// Mitsubishi GX Works2 project: 20国轩1次注液出11.16和条码枪通信   PLC: Q06UDEH (continued)
	
	(*U1任务处理 *)
	m_TPU1TaskComplete(IN:=ConveyorIO20110.xEmpty ,PT:=t#200ms,Q:= m_xU1TaskComplete,ET:= m_tU1TaskComplete );
	(*这里东西运走之后延时200ms再完成任务，这个时间是防止扫描周期的影响，让U型块先复位，再完成任务*)
Task20301(	xCondition:=TaskCondition20301,
 xTaskComplete:=LDF(TRUE,m_xU1TaskComplete),
 xReset:=g_xResetSingle AND g_diDeviceIDSelect=20110,
 iPriority:=UConveyorIO20301.iTask);
	TaskCondition20301[1]:=NOT ConveyorIO20101.xEmpty  AND LifterIO20201.iCurrentPos=2  AND X2F AND m_i20101Task>0;
	TaskCondition20301[2]:=(NOT ConveyorIO201021.xEmpty AND ConveyorIO201021.diDesConveyor=20115) 
												OR(NOT  ConveyorIO20110.xEmpty AND (ConveyorIO20110.diDesConveyor<>20102 OR ConveyorIO20110.diDesConveyor<>20103)) ;
	TaskCondition20301[3]:=(NOT ConveyorIO201031.xEmpty AND ConveyorIO201031.diDesConveyor=20115)
												OR (NOT  ConveyorIO20110.xEmpty AND(ConveyorIO20110.diDesConveyor<>20102 OR ConveyorIO20110.diDesConveyor<>20103));
	(*U2Task	*)
	m_TPU2TaskComplete(IN:=ConveyorIO20111.xEmpty ,PT:=t#200ms,Q:= m_xU2TaskComplete,ET:= m_tU2TaskComplete );
	Task20303(	xCondition:=TaskCondition20303,
 	xTaskComplete:=LDf(TRUE, m_xU2TaskComplete),
 	xReset:=g_xResetSingle AND g_diDeviceIDSelect=20111,
 	iPriority:=UConveyorIO20303.iTask);
		TaskCondition20303[1]:=NOT ConveyorIO20110.xEmpty AND NOT  (ConveyorIO20110.diDesConveyor=20103 
																OR ConveyorIO20110.diDesConveyor=20102
																OR ConveyorIO20110.diDesConveyor=0)(*不去左，不去右，也不是0，就认为可以接料*);
		TaskCondition20303[2]:=(NOT ConveyorIO201041.xEmpty  AND ConveyorIO201041.diDesConveyor=20115) 
													OR (NOT ConveyorIO20111.xEmpty AND (ConveyorIO20111.diDesConveyor<>20103 OR ConveyorIO20111.diDesConveyor<>20102) );
		TaskCondition20303[3]:=(NOT ConveyorIO201051.xEmpty  AND ConveyorIO201051.diDesConveyor=20115) 
													OR (NOT ConveyorIO20111.xEmpty AND (ConveyorIO20111.diDesConveyor<>20103 OR ConveyorIO20111.diDesConveyor<>20102));
	(*//U3Task*)
	m_TPU3TaskComplete(IN:=ConveyorIO20113.xEmpty ,PT:=t#200ms,Q:= m_xU3TaskComplete,ET:= m_tU3TaskComplete );
	Task20305(	xCondition:=TaskCondition20305,
 	xTaskComplete:=LDF(TRUE,m_xU3TaskComplete),
 	xReset:=g_xResetSingle AND g_diDeviceIDSelect=20113,
 	iPriority:=UConveyorIO20305.iTask);
		TaskCondition20305[1]:=NOT ConveyorIO20112.xEmpty(* AND  (ConveyorIO20112.diDesConveyor=20104 
																OR ConveyorIO20112.diDesConveyor=20105
																OR ConveyorIO20112.diDesConveyor=0);(*不去左，不去右，也不是0，就认为可以接料*) ;
		TaskCondition20305[2]:=(NOT ConveyorIO201061.xEmpty AND ConveyorIO201061.diDesConveyor=20115) 
													OR (NOT ConveyorIO20113.xEmpty AND (ConveyorIO20113.diDesConveyor<>20104 OR ConveyorIO20113.diDesConveyor<>20105));
		TaskCondition20305[3]:=(NOT ConveyorIO201071.xEmpty AND ConveyorIO201071.diDesConveyor=20115)
													OR (NOT ConveyorIO20113.xEmpty AND  (ConveyorIO20113.diDesConveyor<>20104 OR ConveyorIO20113.diDesConveyor<>20105));
	(*//U4Task*)
	m_TPU4TaskComplete(IN:=ConveyorIO20114.xEmpty ,PT:=t#200ms,Q:= m_xU4TaskComplete,ET:= m_tU4TaskComplete );
	Task20307(	xCondition:=TaskCondition20307,
 	xTaskComplete:=LDF(TRUE, m_xU4TaskComplete),
 	xReset:=g_xResetSingle AND g_diDeviceIDSelect=20114,
 	iPriority:=UConveyorIO20307.iTask);
		TaskCondition20307[1]:=NOT ConveyorIO20113.xEmpty  AND NOT (ConveyorIO20113.diDesConveyor=20106
																OR ConveyorIO20113.diDesConveyor=20107
																OR ConveyorIO20113.diDesConveyor=0)
(*																AND ConveyorIo20115.xEmpty*);		
		TaskCondition20307[3]:=((NOT ConveyorIO201091.xEmpty AND ConveyorIO201091.diDesConveyor=20115)
													OR (NOT ConveyorIO20114.xEmpty AND (ConveyorIO20114.diDesConveyor<>20109 OR ConveyorIO20114.diDesConveyor<>20108) ))
(*													AND ConveyorIo20115.xEmpty*);
		TaskCondition20307[2]:=((NOT ConveyorIO201081.xEmpty AND ConveyorIO201081.diDesConveyor=20115)
													OR (NOT ConveyorIO20114.xEmpty AND (ConveyorIO20114.diDesConveyor<>20109 OR ConveyorIO20114.diDesConveyor<>20108) ))
(*													AND ConveyorIo20115.xEmpty*);
(*目标地址的传递，横纵分开传递*)
	ConveyorIO20110.diDesConveyorIn:=	ConveyorIO20101.diDesConveyorOut;
	ConveyorIO20111.diDesConveyorIn:=	ConveyorIO20110.diDesConveyorOut;
	ConveyorIO20112.diDesConveyorIn:=	ConveyorIO20111.diDesConveyorOut;
	ConveyorIO20113.diDesConveyorIn:=	ConveyorIO20112.diDesConveyorOut;
	ConveyorIO20114.diDesConveyorIn:=	ConveyorIO20113.diDesConveyorOut;		
(*纵向传递*)
	ConveyorIO20102.diDesConveyorIn:=	ConveyorIO201021.diDesConveyorOut;
	ConveyorIO20103.diDesConveyorIn:=	ConveyorIO201031.diDesConveyorOut;
	ConveyorIO20104.diDesConveyorIn:=	ConveyorIO201041.diDesConveyorOut;
	ConveyorIO20105.diDesConveyorIn:=	ConveyorIO201051.diDesConveyorOut;
	ConveyorIO20106.diDesConveyorIn:=	ConveyorIO201061.diDesConveyorOut;
	ConveyorIO20107.diDesConveyorIn:=	ConveyorIO201071.diDesConveyorOut;
	ConveyorIO20108.diDesConveyorIn:=	ConveyorIO201081.diDesConveyorOut;
	ConveyorIO20109.diDesConveyorIn:=	ConveyorIO201091.diDesConveyorOut;	
	

IF g_xAuto THEN
	D201.0:=ConveyorIO201221.xEmpty;
	Switchio20311.xEntryEnable:=
	D401.0;(*两个PLC通信，以太网方式*)
	Switchio20311.xSwithEnable:=1;
	Switchio20311.xExitEnable:=ConveyorIO201231.xEmpty;
	ConveyorIO201231.xLoad:=ConveyorIO20122.xNextRun;
	ConveyorIO201231.xUnload:=ConveyorIO20123.xEmpty;
	ConveyorIO20123.xLoad:=	ConveyorIO201231.xNextRun;;	
	ConveyorIO20123.xUnload:=	ConveyorIO20124.xEmpty;
	ConveyorIO20124.xLoad:=	ConveyorIO20123.xNextRun;	
	ConveyorIO20124.xUnload:=	ConveyorIO20125.xEmpty;
	SwitchIO20312.xEntryEnable:=ConveyorIO20124.xNextRun;
	SwitchIO20312.xSwithEnable:=1;
	SwitchIO20312.xLiftCylinderExtendInit:=1;
	SwitchIO20312.xExitEnable:=ConveyorIO201261.xEmpty;     
	ConveyorIO201261.xLoad:=ConveyorIO20126.xNextRun;
	ConveyorIO201261.xUnload:=ConveyorIO20127.xEmpty;
	ConveyorIO20127.xLoad:=	ConveyorIO201261.xNextRun;	
	ConveyorIO20127.xUnload:=	ConveyorIO20128.xEmpty;
	ConveyorIO20128.xLoad:=	ConveyorIO20127.xNextRun;	
	ConveyorIO20128.xUnload:=	ConveyorIO20129.xEmpty;
	ConveyorIO20129.xLoad:=	ConveyorIO20128.xNextRun;	
	ConveyorIO20129.xUnload:=	ConveyorIO20130.xEmpty AND NOT ConveyorIO20130.xError;
	ConveyorIO20130.xLoad:=	ConveyorIO20129.xNextRun;	
	ConveyorIO20130.xUnload:=ConveyorIO20101.xEmpty AND LifterIO20201.iCurrentPos=1 AND X2E AND NOT ConveyorIO20101.xError;
	ConveyorIO20101.xLoad:=ConveyorIO20130.xNextRun AND LifterIO20201.iCurrentPos=1 AND X2E;(*运到升降机上了*)
	LifterIO20201.xMDIExe:=NOT 	ConveyorIO20101.xError
													AND NOT ConveyorIO20130.xError
													AND NOT ConveyorIO20110.xError;
	IF ConveyorIO20101.xEmpty THEN
		LifterIO20201.iDestinationPos:=1;
	ELSE
		LifterIO20201.iDestinationPos:=2;
	END_IF;
	m_TonU1TaskStart(IN:=ConveyorIO20110.xEmpty AND UConveyorIO20301.iTask=1  ,PT:= t#1s ,Q:=m_xU1TaskStart,ET:= m_tU1TaskStart );
	ConveyorIO20101.xUnload:=m_xU1TaskStart  AND 
   															LifterIO20201.iCurrentPos=2 AND X2F
 															 (*AND UConveyorIO20301.iTask=1       这个信号会波动
 															 AND ConveyorIO20110.xEmpty*);
 	ConveyorIO20101.xUnloadCCW:=1;
   
	(*//U1*)	
	UConveyorIO20301.xEntryEnable1:= ConveyorIO20101.xNextRun;
	UConveyorIO20301.xEntryEnable2:=ConveyorIO201021.xNextRun;
	UConveyorIO20301.xEntryEnable3:=ConveyorIO201031.xNextRun;
	
	m_TonU2TaskStart(IN:=ConveyorIO20111.xEmpty  ,PT:= t#300ms ,Q:=m_xU2TaskStart,ET:= m_tU2TaskStart );
	UConveyorIO20301.xExitEnable1:= m_xU2TaskStart AND UConveyorIO20303.iTask=1;
	UConveyorIO20301.xExitEnable2:=ConveyorIO201021.xEmpty;
	UConveyorIO20301.xExitEnable3:=ConveyorIO201031.xEmpty;
	(*//U1接料*)
	ConveyorIO201021.xload:=	ConveyorIO20102.xNextRun;
	ConveyorIO201031.xload:=	ConveyorIO20103.xNextRun;
	(*单电控夹紧气缸动作控制*)
	m_xCatchCylinder[2]:=NOT ConveyorIO201021.xEmpty AND ConveyorIO201021.diDesConveyor=0;
	m_xCatchCylinder[3]:=NOT ConveyorIO201031.xEmpty AND ConveyorIO201031.diDesConveyor=0;
	(*//U1出料Unload	*)
		ConveyorIO201021.xUnload:=ConveyorIO20102.xEmpty AND UConveyorIO20301.iTask=2;
		ConveyorIO201031.xUnload:=ConveyorIO20103.xEmpty AND UConveyorIO20301.iTask=3;

	(**//U2*)
	UConveyorIO20303.xEntryEnable1:= ConveyorIO20110.xNextRun ;
	UConveyorIO20303.xEntryEnable2:=ConveyorIO201041.xNextRun;
	UConveyorIO20303.xEntryEnable3:=ConveyorIO201051.xNextRun;
	UConveyorIO20303.xExitEnable1:= ConveyorIO20112.xEmpty;
	UConveyorIO20303.xExitEnable2:=ConveyorIO201041.xEmpty;
	UConveyorIO20303.xExitEnable3:=ConveyorIO201051.xEmpty;
	(*//U2接料	*)
	ConveyorIO201041.xload:=	ConveyorIO20104.xNextRun;
	ConveyorIO201051.xload:=	ConveyorIO20105.xNextRun;
		(*单电控夹紧气缸动作控制*)
	m_xCatchCylinder[4]:=NOT ConveyorIO201041.xEmpty AND ConveyorIO201041.diDesConveyor=0;
	m_xCatchCylinder[5]:=NOT ConveyorIO201051.xEmpty AND ConveyorIO201051.diDesConveyor=0;
	(*//U2出料Unload	*)
		ConveyorIO201041.xUnload:=ConveyorIO20104.xEmpty AND UConveyorIO20303.iTask=2;
		ConveyorIO201051.xUnload:=ConveyorIO20105.xEmpty AND UConveyorIO20303.iTask=3;
	(*//中间传输*)
	ConveyorIO20112.xLoad:=ConveyorIO20111.xNextRun;
	m_TonU3TaskStart(IN:=ConveyorIO20113.xEmpty  ,PT:= t#300ms ,Q:=m_xU3TaskStart,ET:= m_tU3TaskStart );
	ConveyorIO20112.xUnload:=m_xU3TaskStart AND UConveyorIO20305.iTask=1;
	
	(*//U3	*)
	UConveyorIO20305.xEntryEnable1:= ConveyorIO20112.xNextRun;
	UConveyorIO20305.xEntryEnable2:=ConveyorIO201061.xNextRun;
	UConveyorIO20305.xEntryEnable3:=ConveyorIO201071.xNextRun;
	
	m_TonU4TaskStart(IN:=ConveyorIO20114.xEmpty  ,PT:= t#300ms ,Q:=m_xU4TaskStart,ET:= m_tU4TaskStart );
	UConveyorIO20305.xExitEnable1:= m_xU4TaskStart AND UConveyorIO20307.iTask=1 ;
	UConveyorIO20305.xExitEnable2:=ConveyorIO201061.xEmpty;
	UConveyorIO20305.xExitEnable3:=ConveyorIO201071.xEmpty;
	(*	//U3接料*)
	ConveyorIO201061.xload:=	ConveyorIO20106.xNextRun;
	ConveyorIO201071.xload:=	ConveyorIO20107.xNextRun;
		(*单电控夹紧气缸动作控制*)
	m_xCatchCylinder[6]:=NOT ConveyorIO201061.xEmpty AND ConveyorIO201061.diDesConveyor=0;
	m_xCatchCylinder[7]:=NOT ConveyorIO201071.xEmpty AND ConveyorIO201071.diDesConveyor=0;
	(*//U3出料Unload	*)
		ConveyorIO201061.xUnload:=ConveyorIO20106.xEmpty AND  UConveyorIO20305.iTask=2;
		ConveyorIO201071.xUnload:=ConveyorIO20107.xEmpty AND UConveyorIO20305.iTask=3;
	
	(*//U4	*)
	UConveyorIO20307.xEntryEnable1:= ConveyorIO20113.xNextRun ;
	UConveyorIO20307.xEntryEnable2:=ConveyorIO201081.xNextRun;
	UConveyorIO20307.xEntryEnable3:=ConveyorIO201091.xNextRun;
	UConveyorIO20307.xExitEnable1:= ConveyorIO20115.xEmpty ;
	UConveyorIO20307.xExitEnable2:=ConveyorIO201081.xEmpty;
	UConveyorIO20307.xExitEnable3:=ConveyorIO201091.xEmpty;
	(*	//U4接料*)
	ConveyorIO201081.xload:=	ConveyorIO20108.xNextRun;
	ConveyorIO201091.xload:=	ConveyorIO20109.xNextRun;
		(*单电控夹紧气缸动作控制*)
	m_xCatchCylinder[8]:=NOT ConveyorIO201081.xEmpty AND ConveyorIO201081.diDesConveyor=0;
	m_xCatchCylinder[9]:=NOT ConveyorIO201091.xEmpty AND ConveyorIO201091.diDesConveyor=0;
	(*//U4出料Unload	*)
	ConveyorIO201081.xUnload:=ConveyorIO20108.xEmpty AND UConveyorIO20307.iTask=2;
	ConveyorIO201091.xUnload:=ConveyorIO20109.xEmpty AND UConveyorIO20307.iTask=3;
	SwitchIO20309.xEntryEnable:=	ConveyorIO20114.xNextRun;
	SwitchIO20309.xSwithEnable:=1;
	SwitchIO20309.xExitEnable:=ConveyorIO201161.xEmpty;
	ConveyorIO201161.xLoad:=ConveyorIO20116.xNextRun;
	ConveyorIO201161.xUnload:=ConveyorIO20117.xEmpty;
	ConveyorIO20117.xLoad:=ConveyorIO201161.xNextRun;
	ConveyorIO20117.xUnload:=ConveyorIO20118.xEmpty;
	ConveyorIO20118.xLoad:=ConveyorIO20117.xNextRun;
	ConveyorIO20118.xUnload:=ConveyorIO20119.xEmpty AND (g_xScanDone OR SM400);
	Y252:=NOT ConveyorIO20118.xNextRun;
	ConveyorIo20119.tLoadDelay:=T#6s;	
	SwitchIO20310.xEntryEnable:=ConveyorIO20118.xNextRun;
	SwitchIO20310.xLiftCylinderExtendInit:=1;
	SwitchIO20310.xSwithEnable:=1;
	SwitchIO20310.xExitEnable:=D401.2;
	D201.2:=ConveyorIO201191.xNextRun;
(*	ConveyorIO20119.xPutInto:=NOT ConveyorIO20119.xCWPresent AND SM412;
	ConveyorIO201191.xPutInto:=NOT ConveyorIO201191.xCWPresent AND SM412;*)
	(*至此，托盘循环完成*)
	
END_IF;(*g_xAuto那个IF**)	
	(*******************************以下部分为机械手控制*********************************************)
		(*1号机器人*)
		(*位置1*)
		(*发送给机器人的可以放料信号*)
	g_xRobot1Pos1Ready:=NOT ConveyorIO201021.xEmpty   (*线体不为空*)
												AND ConveyorIO201021.diDesConveyor=0(*无目标线体位置*)
												AND NOT g_xRobot1Pos2Ready(*与位置2的信号互锁，同时只有一个ready信号*)
												AND g_xAuto;
		(*接收机器人的完成信号*)
	DMOV(g_xRobot1Pos1Done,20115,ConveyorIO201021.diDesConveyor);(*将目标位置设置成出料线体*)
		(*位置2*)
		(*发送给机器人的可以放料信号*)
	g_xRobot1Pos2Ready:=NOT ConveyorIO201031.xEmpty  (*线体不为空*)
												AND ConveyorIO201031.diDesConveyor=0(*无目标线体位置*)
												AND NOT g_xRobot1Pos1Ready(*与位置1的信号互锁，同时只有一个ready信号*)
												AND g_xAuto;
			(*接收机器人的完成信号*)
	DMOV(g_xRobot1Pos2Done,20115,ConveyorIO201031.diDesConveyor);
	(*2号机器人*)
	g_xRobot2Pos1Ready:=NOT ConveyorIO201041.xEmpty 
												AND ConveyorIO201041.diDesConveyor=0
												AND NOT g_xRobot2Pos2Ready
												AND g_xAuto;
	DMOV(g_xRobot2Pos1Done,20115,ConveyorIO201041.diDesConveyor);
	g_xRobot2Pos2Ready:=NOT ConveyorIO201051.xEmpty 
												AND ConveyorIO201051.diDesConveyor=0
												AND NOT g_xRobot2Pos1Ready 
												AND g_xAuto;
	DMOV(g_xRobot2Pos2Done,20115,ConveyorIO201051.diDesConveyor);
			(*3号机器人*)
		(*位置1*)
		(*发送给机器人的可以放料信号*)
	g_xRobot3Pos1Ready:=NOT ConveyorIO201061.xEmpty   (*线体不为空*)
												AND ConveyorIO201061.diDesConveyor=0(*无目标线体位置*)
												AND NOT g_xRobot3Pos2Ready(*与位置2的信号互锁，同时只有一个ready信号*)
												AND g_xAuto;
		(*接收机器人的完成信号*)
	DMOV(g_xRobot3Pos1Done,20115,ConveyorIO201061.diDesConveyor);(*将目标位置设置成出料线体*)
		(*位置2*)
		(*发送给机器人的可以放料信号*)
	g_xRobot3Pos2Ready:=NOT ConveyorIO201071.xEmpty  (*线体不为空*)
												AND ConveyorIO201071.diDesConveyor=0(*无目标线体位置*)
												AND NOT g_xRobot3Pos1Ready(*与位置1的信号互锁，同时只有一个ready信号*) 
												AND g_xAuto;
			(*接收机器人的完成信号*)
	DMOV(g_xRobot3Pos2Done,20115,ConveyorIO201071.diDesConveyor);
			(*4号机器人*)
		(*位置1*)
		(*发送给机器人的可以放料信号*)
	g_xRobot4Pos1Ready:=NOT ConveyorIO201081.xEmpty   (*线体不为空*)
												AND ConveyorIO201081.diDesConveyor=0(*无目标线体位置*)
												AND NOT g_xRobot4Pos2Ready(*与位置2的信号互锁，同时只有一个ready信号*) 
												AND g_xAuto;
		(*接收机器人的完成信号*)
	DMOV(g_xRobot4Pos1Done,20115,ConveyorIO201081.diDesConveyor);(*将目标位置设置成出料线体*)
		(*位置4*)
		(*发送给机器人的可以放料信号*)
	g_xRobot4Pos2Ready:=NOT ConveyorIO201091.xEmpty  (*线体不为空*)
												AND ConveyorIO201091.diDesConveyor=0(*无目标线体位置*)
												AND NOT g_xRobot4Pos1Ready(*与位置1的信号互锁，同时只有一个ready信号*) 
												AND g_xAuto;
			(*接收机器人的完成信号*)
	DMOV(g_xRobot4Pos2Done,20115,ConveyorIO201091.diDesConveyor);
		
	(*******************************以上部分为机械手控制*********************************************)
	
IF NOT g_xAuto THEN
	D201.0:=0;
	D201.2:=0;
	ConveyorIO201021.diDesConveyor:=0;
	ConveyorIO201031.diDesConveyor:=0;	
	ConveyorIO201041.diDesConveyor:=0;
	ConveyorIO201051.diDesConveyor:=0;
	ConveyorIO201061.diDesConveyor:=0;
	ConveyorIO201071.diDesConveyor:=0;	
	ConveyorIO201081.diDesConveyor:=0;
	ConveyorIO201091.diDesConveyor:=0;	
	g_xRobot1Pos1Ready:=0;
	g_xRobot1Pos2Ready:=0;
	g_xRobot2Pos1Ready:=0;
	g_xRobot2Pos2Ready:=0;
	g_xRobot3Pos1Ready:=0;
	g_xRobot3Pos2Ready:=0;
	g_xRobot4Pos1Ready:=0;
	g_xRobot4Pos2Ready:=0;
	
END_IF;
(*//统计计数*)

ADD_E(LDP(TRUE,NOT ConveyorIO201021.xEmpty)AND UConveyorIO20301.iTask=1,	D10,	1,	D10 );
ADD_E(LDP(TRUE,NOT ConveyorIO201031.xEmpty)AND UConveyorIO20301.iTask=1,	D12,	1,	D12 );
ADD_E(LDP(TRUE,NOT ConveyorIO201041.xEmpty)AND UConveyorIO20303.iTask=1,	D14,	1,	D14 );
ADD_E(LDP(TRUE,NOT ConveyorIO201051.xEmpty)AND UConveyorIO20303.iTask=1,	D16,	1,	D16 );
ADD_E(LDP(TRUE,NOT ConveyorIO201061.xEmpty)AND UConveyorIO20305.iTask=1,	D18,	1,	D18 );
ADD_E(LDP(TRUE,NOT ConveyorIO201071.xEmpty)AND UConveyorIO20305.iTask=1,	D20,	1,	D20 );
ADD_E(LDP(TRUE,NOT ConveyorIO201081.xEmpty)AND UConveyorIO20307.iTask=1,	D22,	1,	D22 );
ADD_E(LDP(TRUE,NOT ConveyorIO201091.xEmpty)AND UConveyorIO20307.iTask=1,	D24,	1,	D24 );
(*//统计数据清零,这些M都是在触摸屏上的数据清零按钮*)
DMOV(	M62,	0,	D10);
DMOV(	M63,	0,	D12 );
DMOV(	M64,	0,	D14 );
DMOV(	M65,	0,	D16 );
DMOV(	M66,	0,	D18 );
DMOV(	M67,	0,	D20 );
DMOV(	M68,	0,	D22 );
DMOV(	M69,	0,	D24 );
(*临时加一些送出按钮，方便操作*)
DMOVP( M42 ,10115 , ConveyorIO201021.diDesConveyor );
DMOVP( M43 ,10115 , ConveyorIO201031.diDesConveyor );
DMOVP( M44 ,10115 , ConveyorIO201041.diDesConveyor );
DMOVP( M45 ,10115 , ConveyorIO201051.diDesConveyor );
DMOVP( M46 ,10115 , ConveyorIO201061.diDesConveyor );
DMOVP( M47 ,10115 , ConveyorIO201071.diDesConveyor );
DMOVP( M48 ,10115 , ConveyorIO201081.diDesConveyor );
DMOVP( M49 ,10115 , ConveyorIO201091.diDesConveyor );

(*报警*)
g_xAlarm:=NOT g_xEStop;
END_PROGRAM

FUNCTION_BLOCK PreemptivePriority
VAR_INPUT
  xCondition : ARRAY [1..13] OF BOOL;  (* 条件1 *)
  xTaskComplete : BOOL;  (* 任务完成 *)
  xReset : BOOL;  (* 复位 *)
END_VAR
VAR
  xOccupy : BOOL;  (* 占用 *)
END_VAR
VAR_OUTPUT
  iPriority : INT;  (* 输出任务号 *)
END_VAR
VAR
  m_tonConditionDelay : TON;
  m_xConditionDelay : BOOL;
  m_tConditionCurrentTime : TIME;
  m_iLastTask : INT;  (* 上次执行的任务 *)
  m_tpLastTaskPulse1 : TP;
  m_tpLastTaskPulse2 : TP;
  m_tpLastTaskPulse3 : TP;
  m_tpLastTaskPulse4 : TP;
  m_tpLastTaskPulse5 : TP;
  m_xLastTaskPulse : ARRAY [1..13] OF BOOL;
  m_tLastTaskPulse : ARRAY [1..13] OF TIME := [13(T#0s)];
  m_tpLastTaskPulse6 : TON;
  ii : INT;
END_VAR
VAR CONSTANT
  CONDITION_QUANTITY : INT := 9;
END_VAR
VAR
  m_tpLastTaskPulse7 : TON;
  m_tpLastTaskPulse8 : TON;
  m_tpLastTaskPulse9 : TON;
  m_tpLastTaskPulse10 : TON;
  m_tpLastTaskPulse11 : TON;
  m_tpLastTaskPulse12 : TON;
  m_tpLastTaskPulse13 : TON;
END_VAR
(*抢占式优先级块
现在满足13个条件的任务进行抢占式优先级排列
条件满足后延时两秒，开始执行任务，
同一任务连续执行优先级下降
需要改造成任意多个
使用于一个入口多个出口的程序，使用抢占式优先级块
*)
IF LDP(TRUE, xTaskComplete) THEN
	xOccupy:=0;
	iPriority:=0;
END_IF;
(*//任务滤波，延时两秒*)
m_tonConditionDelay(IN:=( xCondition[1]
 	OR xCondition[2]
 	OR xCondition[3]
 	OR xCondition[4]
 	OR xCondition[5]
 	OR xCondition[6]
 	OR xCondition[7]
 	OR xCondition[8]
 	OR xCondition[9]
 	OR xCondition[10]
 	OR xCondition[11]
 	OR xCondition[12]
 	OR xCondition[13]
 	)
 	AND iPriority=0,
 PT:= T#1s,
 Q:= m_xConditionDelay ,
 ET:= m_tConditionCurrentTime );		
(*//判断优先级，上个任务与本次任务相同，延时一秒执行*)
m_tpLastTaskPulse1(IN:= xCondition[1]  AND m_iLastTask=1 AND m_xConditionDelay  ,PT:= T#1s,Q:= m_xLastTaskPulse[1],ET:= m_tLastTaskPulse[1] );
m_tpLastTaskPulse2(IN:= xCondition[2]  AND m_iLastTask=2 AND m_xConditionDelay  ,PT:= T#1s,Q:= m_xLastTaskPulse[2],ET:= m_tLastTaskPulse[2] );
m_tpLastTaskPulse3(IN:= xCondition[3]  AND m_iLastTask=3 AND m_xConditionDelay  ,PT:= T#1s,Q:= m_xLastTaskPulse[3],ET:= m_tLastTaskPulse[3] );
m_tpLastTaskPulse4(IN:= xCondition[4]  AND m_iLastTask=4 AND m_xConditionDelay  ,PT:= T#1s,Q:= m_xLastTaskPulse[4],ET:= m_tLastTaskPulse[4] );
m_tpLastTaskPulse5(IN:= xCondition[5]  AND m_iLastTask=5 AND m_xConditionDelay  ,PT:= T#1s,Q:= m_xLastTaskPulse[5],ET:= m_tLastTaskPulse[5] );
m_tpLastTaskPulse6(IN:= xCondition[6]  AND m_iLastTask=6 AND m_xConditionDelay  ,PT:= T#1s,Q:= m_xLastTaskPulse[6],ET:= m_tLastTaskPulse[6] );
m_tpLastTaskPulse7(IN:= xCondition[7]  AND m_iLastTask=7 AND m_xConditionDelay  ,PT:= T#1s,Q:= m_xLastTaskPulse[7],ET:= m_tLastTaskPulse[7] );
m_tpLastTaskPulse8(IN:= xCondition[8]  AND m_iLastTask=8 AND m_xConditionDelay  ,PT:= T#1s,Q:= m_xLastTaskPulse[8],ET:= m_tLastTaskPulse[8] );
m_tpLastTaskPulse9(IN:= xCondition[9]  AND m_iLastTask=9 AND m_xConditionDelay  ,PT:= T#1s,Q:= m_xLastTaskPulse[9],ET:= m_tLastTaskPulse[9] );
m_tpLastTaskPulse10(IN:= xCondition[10]  AND m_iLastTask=10 AND m_xConditionDelay  ,PT:= T#1s,Q:= m_xLastTaskPulse[10],ET:= m_tLastTaskPulse[10] );
m_tpLastTaskPulse11(IN:= xCondition[11]  AND m_iLastTask=11 AND m_xConditionDelay  ,PT:= T#1s,Q:= m_xLastTaskPulse[11],ET:= m_tLastTaskPulse[11] );
m_tpLastTaskPulse12(IN:= xCondition[12]  AND m_iLastTask=12 AND m_xConditionDelay  ,PT:= T#1s,Q:= m_xLastTaskPulse[12],ET:= m_tLastTaskPulse[12] );
m_tpLastTaskPulse13(IN:= xCondition[13]  AND m_iLastTask=13 AND m_xConditionDelay  ,PT:= T#1s,Q:= m_xLastTaskPulse[13],ET:= m_tLastTaskPulse[13] );
(*//执行*)
FOR ii:=1 TO CONDITION_QUANTITY BY 1 DO 
	IF NOT xCondition[ii] AND NOT xOccupy THEN
		iPriority:=0;
	END_IF;
	IF xCondition[ii] AND NOT xOccupy AND m_xConditionDelay AND NOT  m_xLastTaskPulse[ii]  THEN
		iPriority:=ii;
		xOccupy:=1;
		m_iLastTask:=ii;
	END_IF;
END_FOR;        
(*//复位*)
IF xReset THEN
	iPriority:=0;
	xOccupy:=0;
	m_iLastTask:=0;	
END_IF;
(*//清除占用*)
IF iPriority=0 THEN
	xOccupy:=0;
END_IF;
END_FUNCTION_BLOCK

FUNCTION_BLOCK PriorityQueue
VAR_INPUT
  arrxCondition : ARRAY [1..13] OF QueueElement;
  xTaskComplete : BOOL;  (* 任务完成 *)
  xReset : BOOL;  (* 复位 *)
END_VAR
VAR
  xOccupy : BOOL;  (* 占用 *)
END_VAR
VAR_OUTPUT
  iPriority : INT;  (* 输出任务号 *)
END_VAR
VAR
  jj : INT;
END_VAR
VAR CONSTANT
  CONDITION_QUANTITY : INT := 9;
END_VAR
VAR_IN_OUT
  arriTaskStack : ARRAY [0..13] OF INT;
END_VAR
VAR
  ii : INT;
  kk : INT;
  arrxConditionDelay : ARRAY [1..13] OF BOOL;
  arrxConditionEdgeDetect : ARRAY [1..13] OF BOOL;
  arrxDelayEdgeDetect : ARRAY [1..13] OF BOOL;
  arriDelayCounter : ARRAY [1..13] OF INT;
  ll : INT;
  Temp : INT;
  mm : INT;
  nn : INT;
  Temp2 : INT;
  oo : INT;
END_VAR
(****************************************************************************)
(*
一般情况多对一的任务调度采用这个结构，排队通过出口
优先级功能块，存储任意条件的优先级，实现栈功能先入先出，
复位功能还有问题，
出入栈式优先级块，满足条件后入栈，先入先出，在栈尾加载新任务
栈首为当前执行的任务，任务完成使用上升沿触发，触发后栈首元素弹出

复位功能清空堆栈，栈的容量在CONDITION_QUANTITY 设置
增加了结构体，结构体中带有一个条件函数，和一个优先级指示
任务完成后通过凭借优先级来排序，优先级高的条件先执行   优先级排序是从小到大的，数值小的优先级高
防止干扰，增加了任务的1秒的延时
*)

(***************************************************************************)
(*(//入栈*)
FOR ii:=1 TO CONDITION_QUANTITY BY 1 DO
	(*//循环内无法用定时器，改用计数器的形式*)
	IF arrxCondition[ii].xCondition AND SM411 (*//0.2秒的方波信号，如果移植需要修改成两个定时器*)
		AND arriDelayCounter[ii]<6  (* //计数为6，5个0.2秒的方波，所以为1秒*)
		AND NOT arrxDelayEdgeDetect[ii] THEN    (*//循环内无法用沿函数，增加锁定标志位*)
		arriDelayCounter[ii]:=arriDelayCounter[ii]+1;   (*//计数*)
	END_IF;
	IF NOT arrxCondition[ii].xCondition THEN
		arriDelayCounter[ii]:=0;   (*//计数清零*)
	END_IF;
	arrxDelayEdgeDetect[ii]:=arrxCondition[ii].xCondition AND SM411;  (*//沿函数锁*)
	IF arriDelayCounter[ii]=5 AND NOT arrxConditionEdgeDetect[ii] THEN;  (*//条件满足1秒后*)
		FOR kk:=0 TO CONDITION_QUANTITY BY 1 DO    
			IF arriTaskStack[kk]=0 THEN
				arriTaskStack[kk]:=ii;   (*//栈尾添加*)
				EXIT;
			END_IF;		
		END_FOR;
	END_IF;	
	arrxConditionEdgeDetect[ii]:=arriDelayCounter[ii]=5;  (*//边沿*)
END_FOR;
(*//栈顶任务为当前执行的任务**)
iPriority:=arriTaskStack[0]; 
(*//栈顶任务完成，弹出*)
IF 	LDP(TRUE, xTaskComplete) THEN
	FOR jj:=0 TO CONDITION_QUANTITY-1 BY 1 DO
		arriTaskStack[jj]:=arriTaskStack[jj+1];
	END_FOR;
	arriTaskStack[CONDITION_QUANTITY]:=0;(*//栈尾清零*)
	(*//排序，使用插入排序*)
	FOR oo:=0 TO CONDITION_QUANTITY BY 1 DO
		IF arriTaskStack[oo]=0 THEN
			EXIT;  (* //寻找栈中不为零的元素  ，防止0元素进入条件查找的时候报错*)
		END_IF;
	END_FOR;
	(*//插入排序insertionsort*)
	FOR mm:=1 TO oo-1  BY 1 DO   (*//从1开始*)
		Temp:=arriTaskStack[mm];  (*//当前数据记录 *)
		Temp2:=arrxCondition[arriTaskStack[mm]].iPriority;  (*//当前优先级记录 *)
		nn:=mm;  (*//指针赋值*)
		WHILE  (nn>0 AND Temp2< arrxCondition[arriTaskStack[nn-1]].iPriority)  DO  (*//优先级比较，当前优先级小于他前面元素优先级的时候*)
			 arriTaskStack[nn] := arriTaskStack[nn-1] ;  (*//优先级低的向后复制，比TEMP2大的元素都要复制到下一个位置*)
			 nn:=nn-1;
		END_WHILE;
		arriTaskStack[nn]:=Temp; (*//把当前数据放在合适的位置*)
	END_FOR;
END_IF;
(*//复位*)
IF xReset THEN
	FOR jj:=0 TO CONDITION_QUANTITY BY 1 DO
		arriTaskStack[jj]:=0;
	END_FOR;
	FOR ll:=1 TO CONDITION_QUANTITY BY 1 DO
		arrxConditionEdgeDetect[ll]:=0;
		arriDelayCounter[ll]:=0;
	END_FOR;
END_IF;
END_FUNCTION_BLOCK

FUNCTION_BLOCK ShuttleCar
VAR_IN_OUT
  ShuttleCarInOut : ShuttleCarIO;
END_VAR
VAR
  m_tonBrakeDelay : TON;  (* 延时 *)
  m_tBrakeDelayCurrentTime : TIME;
  m_tonArriveDelay : TON;  (* 到达延时计时器 *)
  m_xArriveDelay : BOOL;  (* 到达延时 *)
  m_tArriveDelayCurrentTime : TIME;  (* 到达延时当前时间 *)
  m_xInit : BOOL;  (* 初始化标志位 *)
  m_tonPauseDelay : TON;  (* 暂停减速 *)
  m_tPauseDelayCurrentTime : TIME;  (* 暂停延时当前时间 *)
  m_tonOvertimeAlarm : TON;  (* 超时报警定时器 *)
  m_tOvertimeCurrentTime : TIME;  (* 超时报警当前时间 *)
END_VAR
(*******************************************************************
输送小车程序，可用于使用认址片控制位置的输送车程序，可用于控制提升机，
使用了限位捕捉程序防止小车惯性过大冲过限位后继续行走，捕捉程序采用反
转复位，这样设计有弊端可能反转复位后车的位置并没有回到限位以内,当两个
限位同时碰到的时候，会使运料小车进入死锁状态，通过xPassLimit来解开死锁，
可以在触摸屏中使用一个带权限的按钮来进行控制，配合ShuttleCarCurrentPos
函数来计算位置信息
增加自动开始后将当前位置置为零的信号防止设备停在两个位置开关的中间
修改信息  修改后请增加版本
2018-1-22增加到位延时：到位延时时间可以设置，适应双向到位的位置开关，通过调整延时时间让穿梭车停在到位开关的中间
增加气缸控制信号 ShuttleCarInOut.xCylinder
增加抱闸延时 ShuttleCarInOut.tBrakeDelay
增加超时报警 ShuttleCarInOut.xOvertimeAlarm
YAO      V1.0
2018-1-22 YAO V1.1
2018-6-3：增加点动xMoveStep，单体报警复位
接口说明：
输入：
xReady    准备就绪信号，接变频器的准备就绪，无准备就绪信号的设备常置1
xForward   手动 正转
xBackward 手动 反转
iCurrentPos 当前位置信息，由外部函数给出
iDestinationPos  目标位置，自动情况下判断目标位置和当前位置的差，选择前进或后退
xPosLimit 正方向限位  常闭信号
xNegLimit 反方向限位  常闭信号
xMDIExe   自动行走使能
xPassLimit 限位屏蔽
tArriveDelay 到位延时时间设置，当前位置等于目标位置后延时相应时间后停止，默认为0
xCylinder 如果是气缸的把这个标志位置为1，
tBrakeDelay 打开抱闸延时，默认100ms。行走后会延时相应的时间打开抱闸，防止提升轴的掉落
xLooseDetect 松绳检测开关
输出：
xCW 正转输出
xCCW 反转输出
xBrake 抱闸输出 
xMDIDone 自动行走完成信号
xPosLimitCatch 正限位报警
xNegLimitCatch 负限位报警
xBusy 工作中信号
xLooseAlarm 松绳报警，报警后不可以下降，提升后如果没有松绳检测开关后复位报警信号


********************************************************************)
IF NOT m_xInit THEN
	ShuttleCarInOut.tArriveDelay:=T#0s;   (*到位延时初始化为0*)
	ShuttleCarInOut.tBrakeDelay:=T#100ms;(*抱闸延时初始化为100ms*)
	ShuttleCarInOut.tSetOverTime:=T#60s;(*超时报警初始化为1分钟*)
	m_xInit:=1;
END_IF;
(*如果是气缸的话屏蔽限位和Ready信号*)
IF ShuttleCarInOut.xCylinder THEN
	ShuttleCarInOut.xPosLimit:=1;
	ShuttleCarInOut.xNegLimit:=1;
	ShuttleCarInOut.xReady:=1;
END_IF;
(*限位捕捉，防止冲过限位开关，反转后复位*)
ShuttleCarInOut.xPosLimitCatch:=LDF(TRUE,ShuttleCarInOut.xPosLimit) OR ShuttleCarInOut.xPosLimitCatch;
IF ShuttleCarInOut.xCCW THEN  
	ShuttleCarInOut.xPosLimitCatch:=0;
END_IF;

ShuttleCarInOut.xNegLimitCatch:=LDF(TRUE,ShuttleCarInOut.xNegLimit) OR ShuttleCarInOut.xNegLimitCatch;
(*松绳报警*)
IF LDP(TRUE,ShuttleCarInOut.xLooseDetect) THEN	
	ShuttleCarInOut.xLooseAlarm:=1;
END_IF;
(*提升复位报警*)
IF ShuttleCarInOut.xCW AND NOT  ShuttleCarInOut.xLooseDetect THEN   
	ShuttleCarInOut.xLooseAlarm:=0; 
END_IF;

IF ShuttleCarInOut.xCW THEN   
	ShuttleCarInOut.xNegLimitCatch:=0; 
END_IF;

IF ShuttleCarInOut.xPassLimit OR
	g_xReset OR   (*增加复位按钮*)
	(ShuttleCarInOut.xNegLimitCatch 
	AND ShuttleCarInOut.xPosLimitCatch)  THEN  
	ShuttleCarInOut.xNegLimitCatch:=0; 
	ShuttleCarInOut.xPosLimitCatch:=0;
	ShuttleCarInOut.xLooseAlarm:=0;
END_IF;
IF ShuttleCarInOut.xReady AND g_xEStop THEN
(*手动*)
    IF g_xManual THEN  
	    IF ShuttleCarInOut.xForward 
			AND ShuttleCarInOut.xBackward=0 
			AND ShuttleCarInOut.xCCW=0 
			AND ShuttleCarInOut.xPosLimitCatch=0  THEN
		    ShuttleCarInOut.xCW:=1;
		    ELSE
		    ShuttleCarInOut.xCW:=0;
	    END_IF;
	    IF ShuttleCarInOut.xBackward 
			AND ShuttleCarInOut.xForward=0 
			AND ShuttleCarInOut.xCW=0 
			AND ShuttleCarInOut.xNegLimitCatch=0 
			AND ShuttleCarInOut.xLooseAlarm=0
			AND G_xEStop THEN  
		    ShuttleCarInOut.xCCW:=1;
		    ELSE
		    ShuttleCarInOut.xCCW:=0;
	    END_IF;
    END_IF;
    (**********)
(*自动*)
  IF g_xAuto OR ShuttleCarInOut.xMoveStep   THEN  
  	(*点动*)
  	IF LDP(TRUE,ShuttleCarInOut.xMoveStep)  THEN (*点动模式后把当前位置赋值给目标位置，防止误动作*)
  		ShuttleCarInOut.iDestinationPos:=ShuttleCarInOut.iCurrentPos;
  		END_IF;
 		IF LDP(TRUE,ShuttleCarInOut.xForward) AND ShuttleCarInOut.xMoveStep THEN
 			ShuttleCarInOut.xMDIExe:=1;
			ShuttleCarInOut.iDestinationPos:=ShuttleCarInOut.iCurrentPos+1;
		END_IF;
		IF LDP(TRUE,ShuttleCarInOut.xBackward) AND ShuttleCarInOut.xMoveStep AND ShuttleCarInOut.iCurrentPos>0  THEN
			ShuttleCarInOut.xMDIExe:=1;
			ShuttleCarInOut.iDestinationPos:=ShuttleCarInOut.iCurrentPos-1;
		END_IF;	 
	(*>>>>>>>>>>>>>>>>>>>>>>>>>>>>>>>>>>>>>*)	
	  IF ShuttleCarInOut.xMDIExe AND ShuttleCarInOut.iDestinationPos<>0 THEN	
	    IF ShuttleCarInOut.iCurrentPos<ShuttleCarInOut.iDestinationPos AND ShuttleCarInOut.xPosLimitCatch=0 THEN   (*正转*)
			ShuttleCarInOut.xCW:=1;
			ShuttleCarInOut.xCCW:=0;
			ShuttleCarInOut.xMDIDone:=0;
		END_IF;

		IF ShuttleCarInOut.iCurrentPos>ShuttleCarInOut.iDestinationPos AND ShuttleCarInOut.xNegLimitCatch=0 AND ShuttleCarInOut.xLooseAlarm=0 THEN   (*反转*)
			ShuttleCarInOut.xCCW:=1;
			ShuttleCarInOut.xCW:=0;
			ShuttleCarInOut.xMDIDone:=0;
		END_IF;
	m_tonArriveDelay(IN:= ShuttleCarInOut.iCurrentPos=ShuttleCarInOut.iDestinationPos ,
	                                    PT:= ShuttleCarInOut.tArriveDelay ,
	                                    Q:= m_xArriveDelay ,
	                                    ET:= m_tArriveDelayCurrentTime);
	     (*到位延时时间可以设置，适应双向到位的位置开关，通过调整延时时间让穿梭车停在到位开关的中间*)
		IF m_xArriveDelay AND NOT ShuttleCarInOut.xCylinder THEN
			ShuttleCarInOut.xCW:=0;
			ShuttleCarInOut.xCCW:=0;
			ShuttleCarInOut.xMDIDone:=1;
			ELSE
			ShuttleCarInOut.xMDIDone:=0;
		END_IF;

		IF ShuttleCarInOut.xPosLimitCatch THEN
			ShuttleCarInOut.xCW:=0;
			ShuttleCarInOut.xMDIDone:=0;
		END_IF;

		IF ShuttleCarInOut.xNegLimitCatch  OR ShuttleCarInOut.xLooseAlarm THEN
			ShuttleCarInOut.xCCW:=0;
			ShuttleCarInOut.xMDIDone:=0;
		END_IF;
		ELSE
		ShuttleCarInOut.xCW:=0;
		ShuttleCarInOut.xCCW:=0;
		ShuttleCarInOut.xMDIDone:=0;
	  END_IF;
	END_IF;
	ELSE  (*无就绪信号   或急停的情况下*)
		ShuttleCarInOut.xCW:=0;
		ShuttleCarInOut.xCCW:=0;	
END_IF;
    (*抱闸延时*)
m_tonBrakeDelay(IN:= ShuttleCarInOut.xCW OR ShuttleCarInOut.xCCW,
                                    PT:= ShuttleCarInOut.tBrakeDelay,
                                    Q:=ShuttleCarInOut.xBrake ,
                                    ET:= m_tBrakeDelayCurrentTime);

(*自动上电后把当前位置清零，防止穿梭车不在开关位置*)
IF LDP(TRUE,g_xAuto) THEN
	ShuttleCarInOut.iCurrentPos:=0;
END_IF;
IF ShuttleCarInOut.xCW OR ShuttleCarInOut.xCCW THEN
	ShuttleCarInOut.xBusy:=1;
	ELSE
	ShuttleCarInout.xBusy:=0;
END_IF;

(*暂停，带延时减速斜坡，ShuttleCarInOut.xPauseRamp为减速斜坡输出位*)
m_tonPauseDelay(IN:=g_xPause,PT:= T#2s ,Q:=ShuttleCarInOut.xPauseRamp,ET:= m_tPauseDelayCurrentTime );
IF ShuttleCarInOut.xPauseRamp THEN
	ShuttleCarInOut.xCW:=0;
	ShuttleCarInOut.xCCW:=0;
	ShuttleCarInOut.xBrake:=0;
END_IF;
(*超时报警*)
m_tonOvertimeAlarm(IN:= ShuttleCarInOut.xMDIExe AND (ShuttleCarInOut.iCurrentPos<>ShuttleCarInOut.iDestinationPos) ,
                                           PT:= ShuttleCarInOut.tSetOverTime,
                                           Q:= ShuttleCarInOut.xOvertimeAlarm ,
                                           ET:= m_tOvertimeCurrentTime );
(*//单体复位，当设备号与本设备一致的时候执行复位*)
IF (g_xResetSingle AND ShuttleCarInOut.diDeviceID=g_diDeviceIDSelect)THEN(*增加单体复位*)
	ShuttleCarInOut.iCurrentPos:=0;
END_IF;
END_FUNCTION_BLOCK

FUNCTION ShuttleCarCurrentPosition
VAR_INPUT
  xPosition1 : BOOL;
  xPosition2 : BOOL;
  xPosition3 : BOOL;
END_VAR
(*//计算输送车当前位置的函数*)
IF xPosition1 THEN
	ShuttleCarCurrentPosition:=1;
END_IF;
IF xPosition2 THEN
	ShuttleCarCurrentPosition:=2;
END_IF;
IF xPosition3 THEN
	ShuttleCarCurrentPosition:=3;
END_IF;
END_FUNCTION

FUNCTION_BLOCK Switch
VAR_IN_OUT
  ConveyorEntryIO : ConveyorIO;
  ConveyorExitIO : ConveyorIO;
END_VAR
VAR
  m_tonLiftCylinderDelay : TON;  (* 顶升延时 *)
  m_xLiftCylinderDelay : BOOL;
  m_tLiftCylinderDelay : TIME;
  m_tonExitBarDelay : TON;  (* 退出阻挡器延时 *)
  m_tExitBarDelay : TIME;
  m_xExitBarDelay : BOOL;
END_VAR
VAR_IN_OUT
  SwitchIO : SwitchIO;
END_VAR
VAR
  iStep : INT;
  m_xInitial : BOOL;
  m_tonCylinderOvertime : TON;  (* 气缸超时报警定时器 *)
  m_tCylinderOvertimeCurrent : TIME;
END_VAR
(**************************************************
//顶升移载模块，抽象为一条输入输线 ，一条输出输送线
//一个进入阻挡器，一个放出阻挡器，和一个顶升气缸的控制
//程序思路比较混乱，接口不清晰，需要整改
//直接放行的时候有问题
//switchEnable =0的时候   离开线体的PutInto有问题
//增加xPutInto程序
//12-17日   V1.0
//***************************************************)
(*ConveyorEntry(ConveyorMotor:=ConveyorEntryIO);
(*ConveyorExit(ConveyorMotor:=ConveyorExitIO);*)


IF NOT m_xInitial THEN
	SwitchIO.tSetOvertime:=T#5s;
	SwitchIO.xExitEnable:=1;
	m_xInitial:=1;
END_IF;
IF g_xAuto THEN
	CASE iStep OF
		0:(*初始化*)
		ConveyorEntryIO.xLoad:=0;
		ConveyorEntryIO.xUnload:=0;
		ConveyorEntryIO.xPutInto:=0;
		ConveyorExitIO.xLoad:=0;
		ConveyorExitIo.xUnload:=0;
		ConveyorExitIO.xPutInto:=0;
		SwitchIO.xEntryBarCylinderRetract:=0;
		SwitchIO.xExitBarCylinderRetract:=0;
		IF SwitchIO.xLiftCylinderExtendInit THEN
			SwitchIO.xLiftCylinderExtend:=1;
			SwitchIO.xLiftCylinderRetract:=0;
		    IF SwitchIO.xLiftCylinderExtendDetect THEN
			    iStep:=1;
			END_IF; 
			ELSE
			SwitchIO.xLiftCylinderExtend:=0;
			SwitchIO.xLiftCylinderRetract:=1;	
		    IF SwitchIO.xLiftCylinderRetractDetect THEN
			    iStep:=1;
		    END_IF;		
		END_IF;
		1:(*上料*)
        IF SwitchIO.xEntryEnable AND ConveyorEntryIO.xEmpty AND ConveyorExitIO.xEmpty THEN
        	SwitchIO.xEntryBarCylinderRetract:=1;
        	ConveyorEntryIO.xLoad:=1;
        END_IF;
        IF ConveyorEntryIO.xEmpty=0 THEN
        	SwitchIO.xEntryBarCylinderRetract:=0;
        	ConveyorEntryIO.xLoad:=0;
        	ConveyorExitIO.xPutInto:=1;
        END_IF;
        IF m_xLiftCylinderDelay AND  SwitchIO.xSwithEnable AND SwitchIO.xExitEnable THEN
			iStep:=2;
        END_IF;
        IF SwitchIO.xSwithEnable=0 AND m_xLiftCylinderDelay AND SwitchIO.xExitEnable  THEN
			iStep:=3;
        END_IF;
		2:(*顶升*)
		ConveyorExitIO.iProductCategory:=ConveyorEntryIO.iProductCategory;
		ConveyorExitIO.iTaskID:=ConveyorEntryIO.iTaskID;
		ConveyorExitIO.diDesConveyor:=ConveyorEntryIO.diDesConveyor;
		SwitchIO.xExitBarCylinderRetract:=0;
		IF SwitchIO.xLiftCylinderExtendInit THEN
			SwitchIO.xLiftCylinderExtend:=0;
			SwitchIO.xLiftCylinderRetract:=1;
		    ELSE
			SwitchIO.xLiftCylinderExtend:=1;
			SwitchIO.xLiftCylinderRetract:=0;			
		END_IF;

		IF SwitchIO.xLiftCylinderExtendInit THEN
		  	IF SwitchIO.xLiftCylinderRetractDetect THEN
		  		iStep:=4;
		  	END_IF;
		  	ELSE
		  	IF SwitchIO.xLiftCylinderExtendDetect THEN
				iStep:=4; 
		  	END_IF;
		END_IF;
		3:(*放行*)	
		ConveyorExitIO.iProductCategory:=ConveyorEntryIO.iProductCategory;
		ConveyorExitIO.iTaskID:=ConveyorEntryIO.iTaskID;
		ConveyorExitIO.diDesConveyor:=ConveyorEntryIO.diDesConveyor;
		SwitchIO.xExitBarCylinderRetract:=1;
		ConveyorExitIO.xPutInto:=0;
		iStep:=4;
		4:(*下料*)
		(*通过出料传输线下料*)
		IF SwitchIO.xExitEnable  AND m_xExitBarDelay AND NOT SwitchIO.xExitBarCylinderRetract  THEN		  
		  	ConveyorExitIO.xUnload:=1;
			ELSE
		  	ConveyorExitIO.xUnload:=0;
		END_IF;	
		(*通过进料传输线下料*)
		IF SwitchIO.xExitEnable  AND m_xExitBarDelay  AND SwitchIO.xExitBarCylinderRetract THEN		  
		  	ConveyorEntryIO.xUnload:=1;
			ELSE
		  	ConveyorEntryIO.xUnload:=0;
		END_IF;			    	
		IF (ConveyorExitIO.xEmpty OR ConveyorEntryIO.xEmpty) AND m_xExitBarDelay  THEN
		  	ConveyorExitIO.xPutInto:=1;
		  	ConveyorEntryIO.xPutInto:=1;
			iStep:=0; 
		END_IF;
	END_CASE;
	m_tonLiftCylinderDelay(IN:=NOT ConveyorEntryIO.xEmpty AND iStep=1 ,PT:= T#1S ,Q:= m_xLiftCylinderDelay ,ET:=m_tLiftCylinderDelay );
	m_tonExitBarDelay(IN:=iStep=4 ,PT:= T#1s ,Q:= m_xExitBarDelay ,ET:= m_tExitBarDelay);
END_IF;
(*复位程序*)
IF (g_xResetSingle AND  (g_diDeviceIDSelect=ConveyorEntryIO.diDeviceID OR g_diDeviceIDSelect=ConveyorExitIO.diDeviceID))
	OR LDP(TRUE,SwitchIO.xLiftCylinderExtendInit) 
	OR LDF(TRUE,SwitchIO.xLiftCylinderExtendInit) 
	OR LDP(TRUE,SwitchIO.xPutInto)  THEN
	ConveyorEntryIO.xPutInto:=1;
	ConveyorExitIO.xPutInto:=1;
	iStep:=0;
END_IF;

